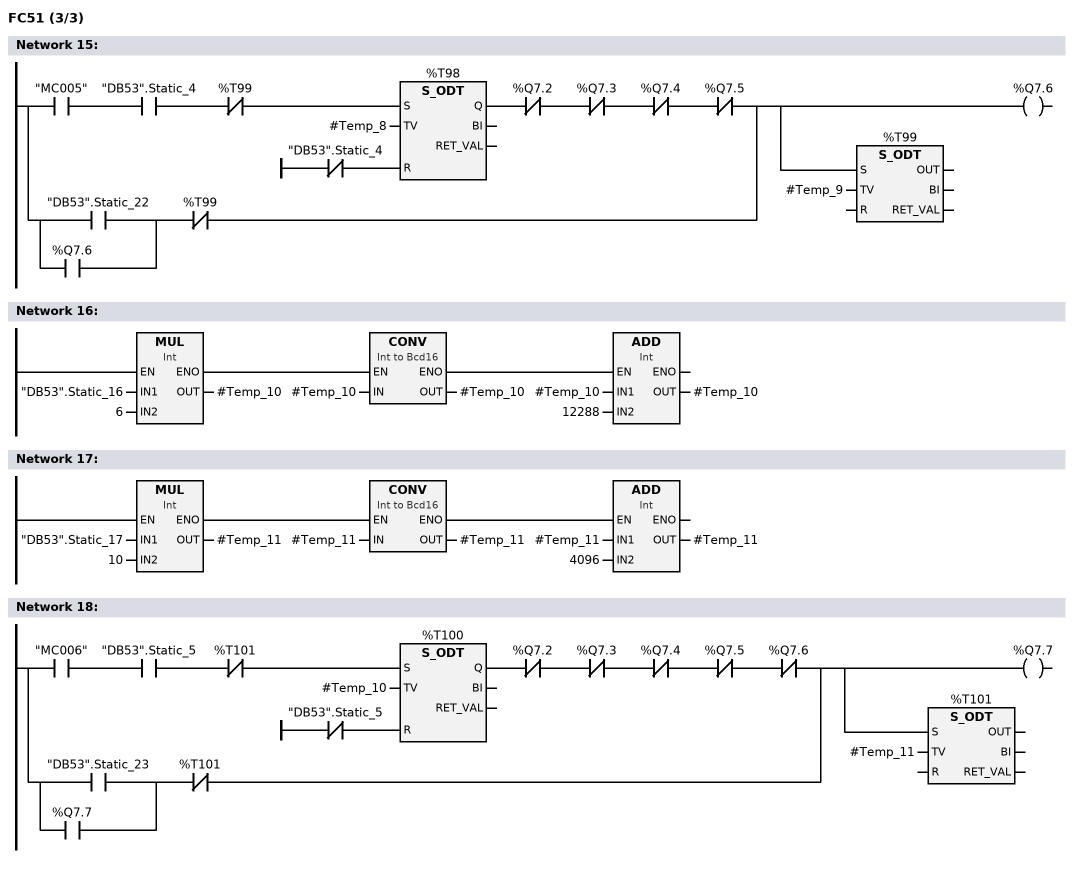
   RUNG wire#powerrail
      Contact( "MC005" )
      Contact( "DB53".Static_4 )
      I_Contact( %T99 )
      S_ODT(T_NO := %T98, TV := #Temp_8, R := wire#w1, BI =>, RET_VAL =>)
      I_Contact( %Q7.2 )
      I_Contact( %Q7.3 )
      I_Contact( %Q7.4 )
      I_Contact( %Q7.5 )
      wire#w2
      Coil( %Q7.6 )
   END_RUNG
   RUNG wire#powerrail
      I_Contact( "DB53".Static_4 )
   END_RUNG wire#w1
   RUNG wire#powerrail
      Contact( "DB53".Static_22 )
      wire#w3
      I_Contact( %T99 )
   END_RUNG wire#w2
   RUNG wire#powerrail
      Contact( %Q7.6 )
   END_RUNG wire#w3
   RUNG wire#w2
      S_ODT(T_NO := %T99, TV := #Temp_9, R :=, BI =>, RET_VAL =>)
   END_RUNG
   // the same network as SCL:
   #_s5time1 := S_ODT(T_NO := %T98,
                      TV := #Temp_8,
                      S := "MC005" AND "DB53".Static_4 AND NOT %T99,
                      R := NOT "DB53".Static_4,
                      Q => #_w1);
   %Q7.6 := (#_w1 AND NOT %Q7.2 AND NOT %Q7.3 AND NOT %Q7.4 AND NOT %Q7.5) OR (("DB53".Static_22 OR %Q7.6) AND NOT %T99);
   #_s5time2 := S_ODT(T_NO := %T99, TV := #Temp_9, S := %Q7.6);
END_REGION

REGION Network 16
   RUNG wire#powerrail
      { S7_Templates := "SrcType := Int"; S7_GenerateENO := "TRUE" } Mul(in1 := "DB53".Static_16, in2 := 6, out => #Temp_10)
      { S7_Templates := "[SrcType := Int, DestType := Bcd16]"; S7_GenerateENO := "TRUE" } Convert(in := #Temp_10, out => #Temp_10)
      { S7_Templates := "SrcType := Int"; S7_GenerateENO := "TRUE" } Add(in1 := #Temp_10, in2 := 12288, out => #Temp_10)
   END_RUNG
   // the same network as SCL:
   // ENO of a box is taken as its EN; it also drops when the box reports an error
   #Temp_10 := "DB53".Static_16 * 6;
   #Temp_10 := INT_TO_BCD16(#Temp_10);
   #Temp_10 := #Temp_10 + 12288;
END_REGION

REGION Network 17
   RUNG wire#powerrail
      { S7_Templates := "SrcType := Int"; S7_GenerateENO := "TRUE" } Mul(in1 := "DB53".Static_17, in2 := 10, out => #Temp_11)
      { S7_Templates := "[SrcType := Int, DestType := Bcd16]"; S7_GenerateENO := "TRUE" } Convert(in := #Temp_11, out => #Temp_11)
      { S7_Templates := "SrcType := Int"; S7_GenerateENO := "TRUE" } Add(in1 := #Temp_11, in2 := 4096, out => #Temp_11)
   END_RUNG
   // the same network as SCL:
   // ENO of a box is taken as its EN; it also drops when the box reports an error
   #Temp_11 := "DB53".Static_17 * 10;
   #Temp_11 := INT_TO_BCD16(#Temp_11);
   #Temp_11 := #Temp_11 + 4096;
END_REGION

REGION Network 18
   RUNG wire#powerrail
      Contact( "MC006" )
      Contact( "DB53".Static_5 )
      I_Contact( %T101 )
      S_ODT(T_NO := %T100, TV := #Temp_10, R := wire#w1, BI =>, RET_VAL =>)
      I_Contact( %Q7.2 )
      I_Contact( %Q7.3 )
      I_Contact( %Q7.4 )
      I_Contact( %Q7.5 )
      I_Contact( %Q7.6 )
      wire#w2
      Coil( %Q7.7 )
   END_RUNG
   RUNG wire#powerrail
      I_Contact( "DB53".Static_5 )
   END_RUNG wire#w1
   RUNG wire#powerrail
      Contact( "DB53".Static_23 )
      wire#w3
      I_Contact( %T101 )
   END_RUNG wire#w2
   RUNG wire#powerrail
      Contact( %Q7.7 )
   END_RUNG wire#w3
   RUNG wire#w2
      S_ODT(T_NO := %T101, TV := #Temp_11, R :=, BI =>, RET_VAL =>)
   END_RUNG
   // the same network as SCL:
   #_s5time1 := S_ODT(T_NO := %T100,
                      TV := #Temp_10,
                      S := "MC006" AND "DB53".Static_5 AND NOT %T101,
                      R := NOT "DB53".Static_5,
                      Q => #_w1);
   %Q7.7 := (#_w1 AND NOT %Q7.2 AND NOT %Q7.3 AND NOT %Q7.4 AND NOT %Q7.5 AND NOT %Q7.6) OR (("DB53".Static_23 OR %Q7.7) AND NOT %T101);
   #_s5time2 := S_ODT(T_NO := %T101, TV := #Temp_11, S := %Q7.7);
END_REGION
END_FUNCTION

ORGANIZATION_BLOCK "Cycle Execution"   // OB1, LAD
{ S7_Optimized_Access := 'FALSE' }
VERSION : 0.1
   VAR_TEMP   // added for the SCL form of the ladder/FBD networks
      _w1 : Bool;
   END_VAR
BEGIN

REGION Network 1
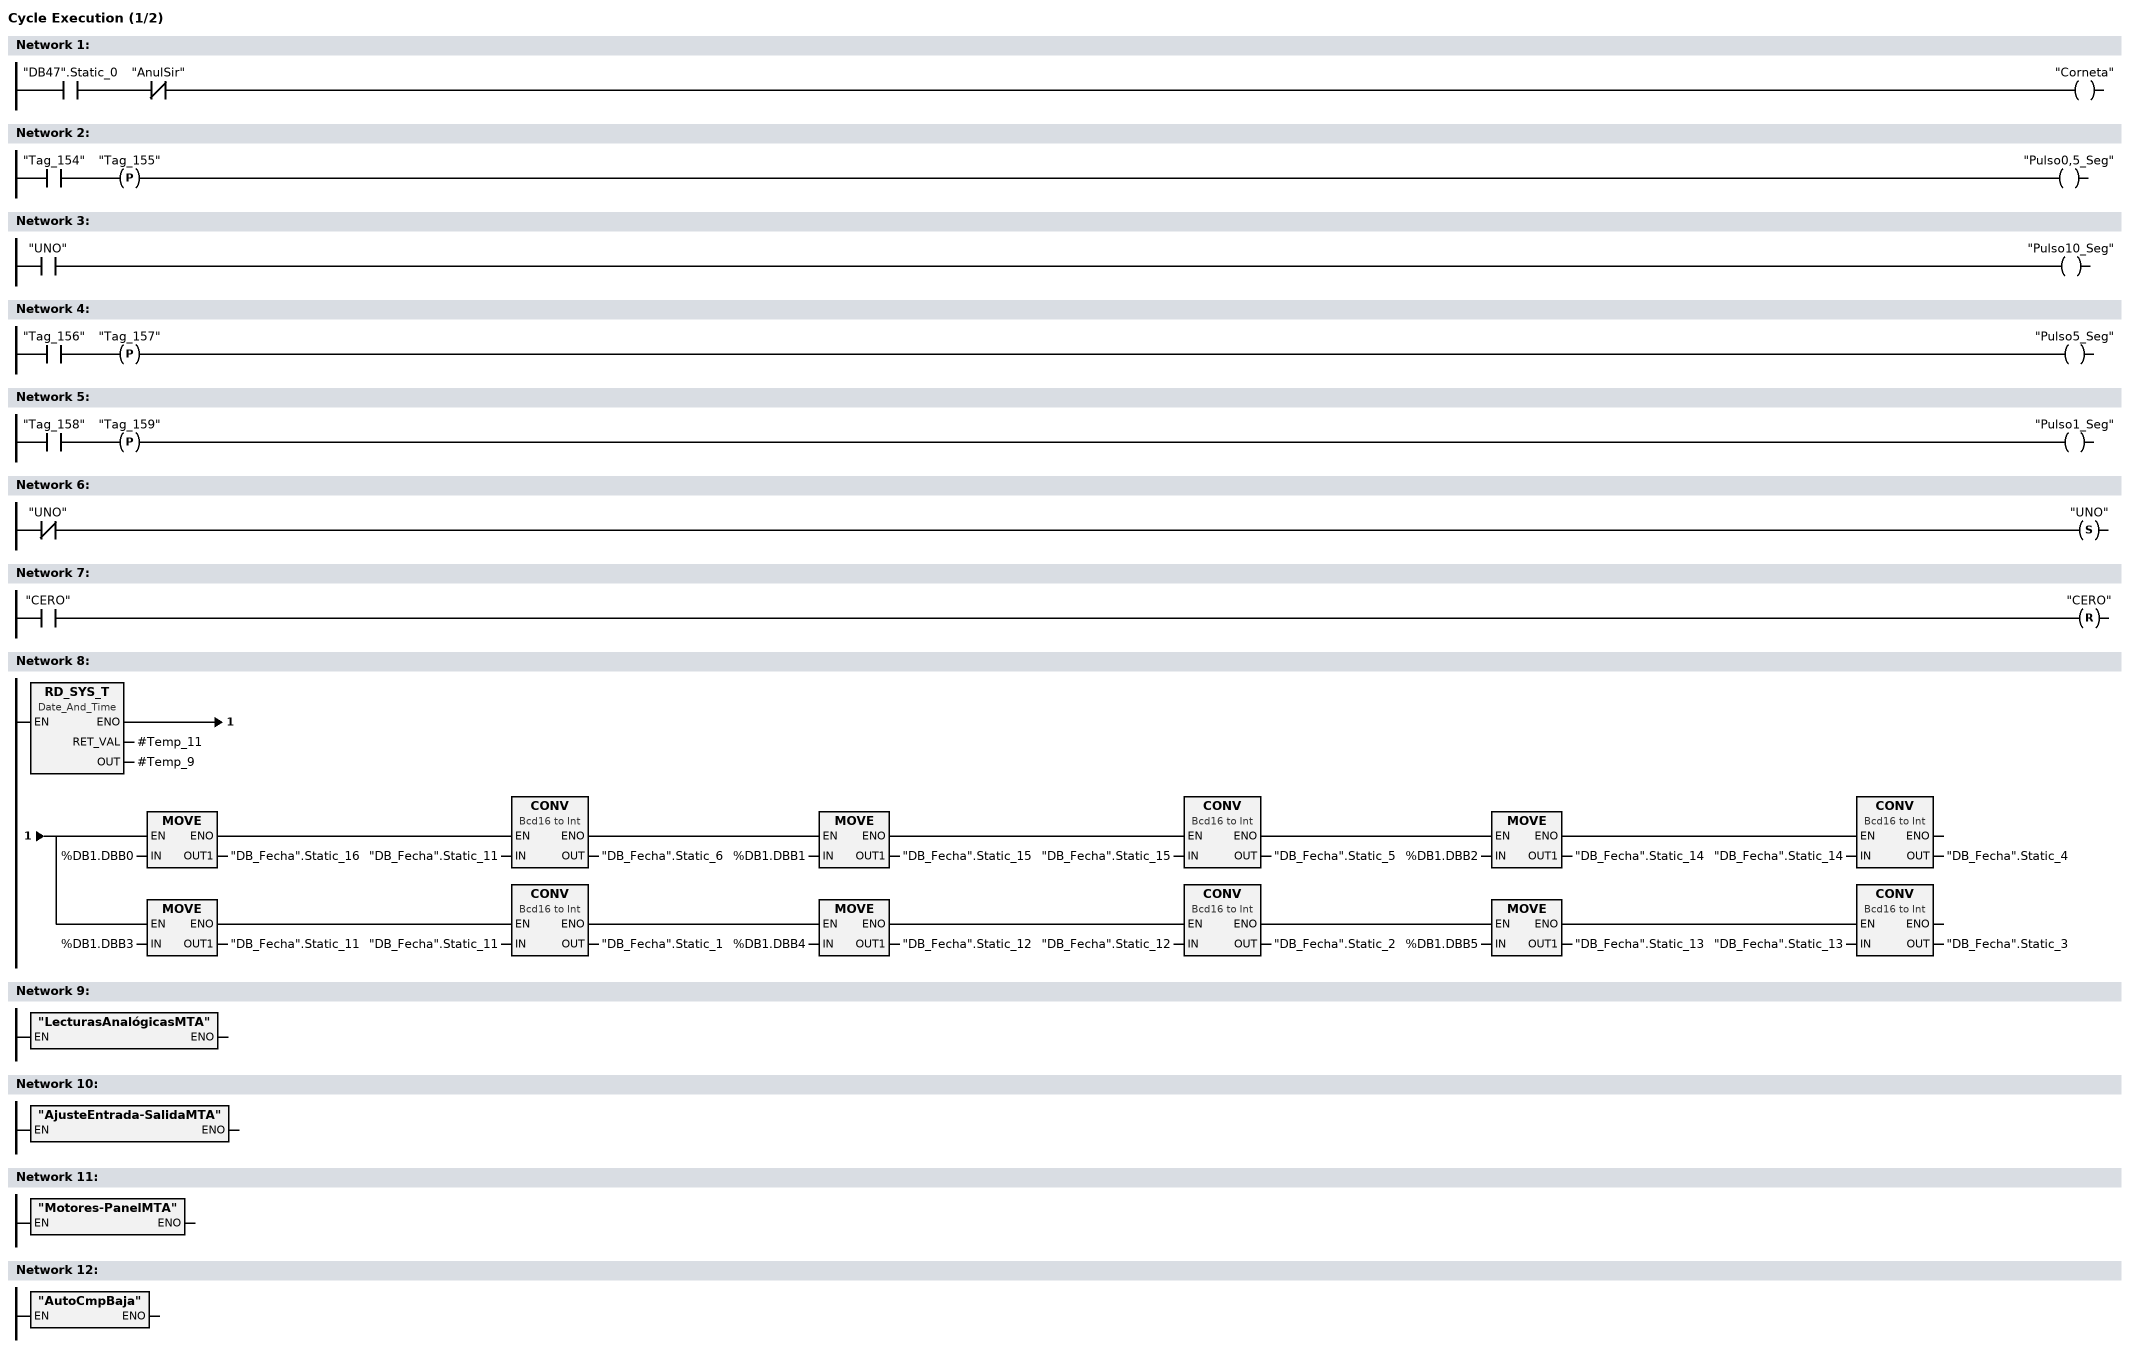
   RUNG wire#powerrail
      Contact( "DB47".Static_0 )
      I_Contact( "AnulSir" )
      Coil( "Corneta" )
   END_RUNG
   // the same network as SCL:
   "Corneta" := "DB47".Static_0 AND NOT "AnulSir";
END_REGION

REGION Network 2
   RUNG wire#powerrail
      Contact( "Tag_154" )
      P_Trig( "Tag_155" )
      Coil( "Pulso0,5_Seg" )
   END_RUNG
   // the same network as SCL:
   #_w1 := "Tag_154" AND NOT "Tag_155";   // rising edge
   "Tag_155" := "Tag_154";
   "Pulso0,5_Seg" := #_w1;
END_REGION

REGION Network 3
   RUNG wire#powerrail
      Contact( "UNO" )
      Coil( "Pulso10_Seg" )
   END_RUNG
   // the same network as SCL:
   "Pulso10_Seg" := "UNO";
END_REGION

REGION Network 4
   RUNG wire#powerrail
      Contact( "Tag_156" )
      P_Trig( "Tag_157" )
      Coil( "Pulso5_Seg" )
   END_RUNG
   // the same network as SCL:
   #_w1 := "Tag_156" AND NOT "Tag_157";   // rising edge
   "Tag_157" := "Tag_156";
   "Pulso5_Seg" := #_w1;
END_REGION

REGION Network 5
   RUNG wire#powerrail
      Contact( "Tag_158" )
      P_Trig( "Tag_159" )
      Coil( "Pulso1_Seg" )
   END_RUNG
   // the same network as SCL:
   #_w1 := "Tag_158" AND NOT "Tag_159";   // rising edge
   "Tag_159" := "Tag_158";
   "Pulso1_Seg" := #_w1;
END_REGION

REGION Network 6
   RUNG wire#powerrail
      I_Contact( "UNO" )
      S_Coil( "UNO" )
   END_RUNG
   // the same network as SCL:
   IF NOT "UNO" THEN "UNO" := TRUE; END_IF;
END_REGION

REGION Network 7
   RUNG wire#powerrail
      Contact( "CERO" )
      R_Coil( "CERO" )
   END_RUNG
   // the same network as SCL:
   IF "CERO" THEN "CERO" := FALSE; END_IF;
END_REGION

REGION Network 8
   // ENO of a box is taken as its EN; it also drops when the box reports an error
   #Temp_11 := RD_SYS_T(out => #Temp_9);
   "DB_Fecha".Static_16 := %DB1.DBB0;
   "DB_Fecha".Static_6 := BCD16_TO_INT("DB_Fecha".Static_11);
   "DB_Fecha".Static_15 := %DB1.DBB1;
   "DB_Fecha".Static_5 := BCD16_TO_INT("DB_Fecha".Static_15);
   "DB_Fecha".Static_14 := %DB1.DBB2;
   "DB_Fecha".Static_4 := BCD16_TO_INT("DB_Fecha".Static_14);
   "DB_Fecha".Static_11 := %DB1.DBB3;
   "DB_Fecha".Static_1 := BCD16_TO_INT("DB_Fecha".Static_11);
   "DB_Fecha".Static_12 := %DB1.DBB4;
   "DB_Fecha".Static_2 := BCD16_TO_INT("DB_Fecha".Static_12);
   "DB_Fecha".Static_13 := %DB1.DBB5;
   "DB_Fecha".Static_3 := BCD16_TO_INT("DB_Fecha".Static_13);
END_REGION

REGION Network 9
   RUNG wire#powerrail
      "LecturasAnalógicasMTA"()
   END_RUNG
   // the same network as SCL:
   "LecturasAnalógicasMTA"();
END_REGION

REGION Network 10
   RUNG wire#powerrail
      "AjusteEntrada-SalidaMTA"()
   END_RUNG
   // the same network as SCL:
   "AjusteEntrada-SalidaMTA"();
END_REGION

REGION Network 11
   RUNG wire#powerrail
      "Motores-PanelMTA"()
   END_RUNG
   // the same network as SCL:
   "Motores-PanelMTA"();
END_REGION

REGION Network 12
   RUNG wire#powerrail
      "AutoCmpBaja"()
   END_RUNG
   // the same network as SCL:
   "AutoCmpBaja"();
END_REGION

REGION Network 13
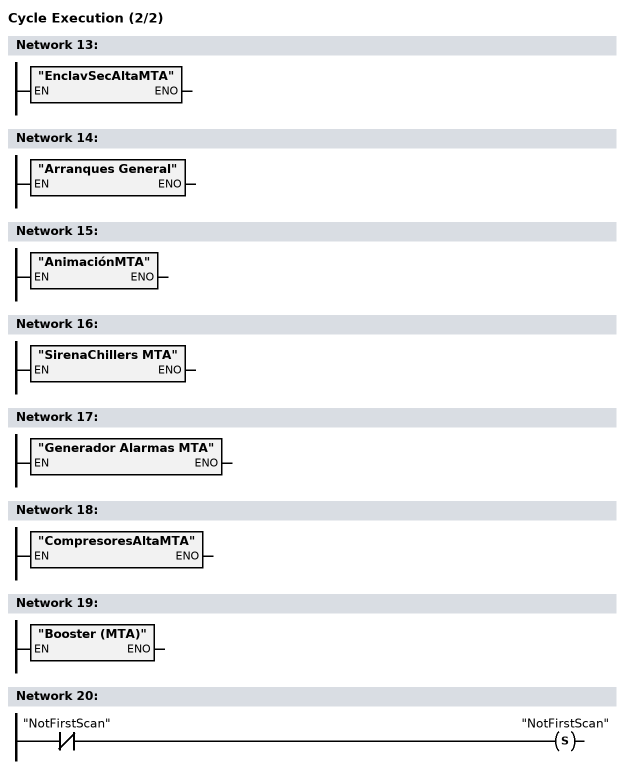
   RUNG wire#powerrail
      "EnclavSecAltaMTA"()
   END_RUNG
   // the same network as SCL:
   "EnclavSecAltaMTA"();
END_REGION

REGION Network 14
   RUNG wire#powerrail
      "Arranques General"()
   END_RUNG
   // the same network as SCL:
   "Arranques General"();
END_REGION

REGION Network 15
   RUNG wire#powerrail
      "AnimaciónMTA"()
   END_RUNG
   // the same network as SCL:
   "AnimaciónMTA"();
END_REGION

REGION Network 16
   RUNG wire#powerrail
      "SirenaChillers MTA"()
   END_RUNG
   // the same network as SCL:
   "SirenaChillers MTA"();
END_REGION

REGION Network 17
   RUNG wire#powerrail
      "Generador Alarmas MTA"()
   END_RUNG
   // the same network as SCL:
   "Generador Alarmas MTA"();
END_REGION

REGION Network 18
   RUNG wire#powerrail
      "CompresoresAltaMTA"()
   END_RUNG
   // the same network as SCL:
   "CompresoresAltaMTA"();
END_REGION

REGION Network 19
   RUNG wire#powerrail
      "Booster (MTA)"()
   END_RUNG
   // the same network as SCL:
   "Booster (MTA)"();
END_REGION

REGION Network 20
   RUNG wire#powerrail
      I_Contact( "NotFirstScan" )
      S_Coil( "NotFirstScan" )
   END_RUNG
   // the same network as SCL:
   IF NOT "NotFirstScan" THEN "NotFirstScan" := TRUE; END_IF;
END_REGION
END_ORGANIZATION_BLOCK

// folder: Alarmas

FUNCTION "SirenaChillers MTA" : Void   // FC7, LAD
{ S7_Optimized_Access := 'FALSE' }
VERSION : 0.1
BEGIN

REGION Network 1
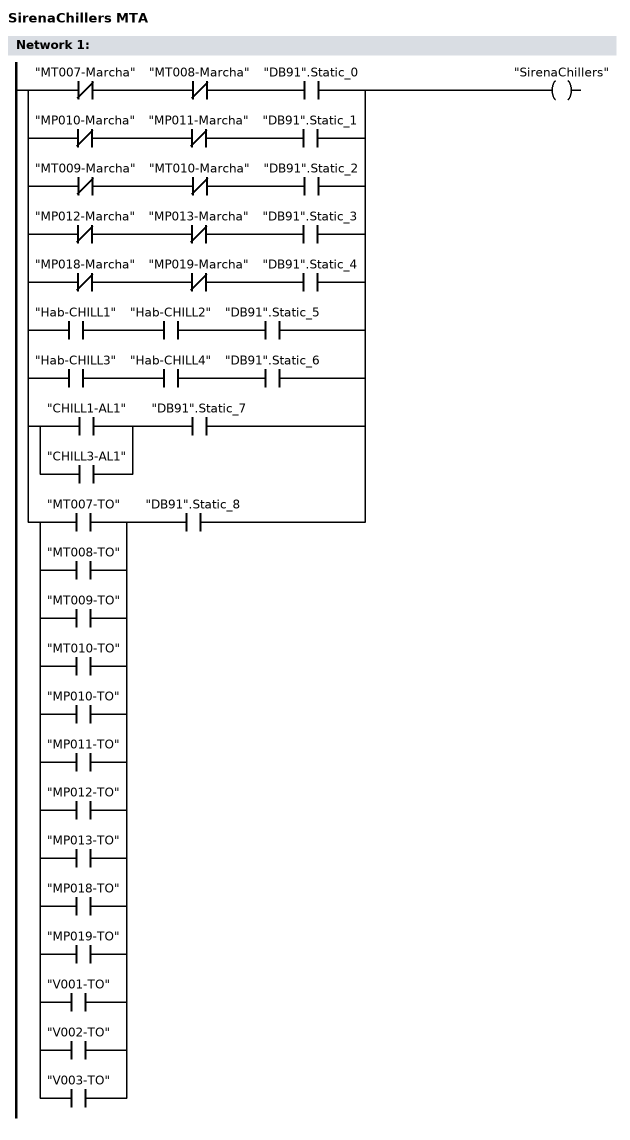
   RUNG wire#powerrail
      I_Contact( "MT007-Marcha" )
      I_Contact( "MT008-Marcha" )
      Contact( "DB91".Static_0 )
      wire#w1
      Coil( "SirenaChillers" )
   END_RUNG
   RUNG wire#powerrail
      I_Contact( "MP010-Marcha" )
      I_Contact( "MP011-Marcha" )
      Contact( "DB91".Static_1 )
   END_RUNG wire#w1
   RUNG wire#powerrail
      I_Contact( "MT009-Marcha" )
      I_Contact( "MT010-Marcha" )
      Contact( "DB91".Static_2 )
   END_RUNG wire#w1
   RUNG wire#powerrail
      I_Contact( "MP012-Marcha" )
      I_Contact( "MP013-Marcha" )
      Contact( "DB91".Static_3 )
   END_RUNG wire#w1
   RUNG wire#powerrail
      I_Contact( "MP018-Marcha" )
      I_Contact( "MP019-Marcha" )
      Contact( "DB91".Static_4 )
   END_RUNG wire#w1
   RUNG wire#powerrail
      Contact( "Hab-CHILL1" )
      Contact( "Hab-CHILL2" )
      Contact( "DB91".Static_5 )
   END_RUNG wire#w1
   RUNG wire#powerrail
      Contact( "Hab-CHILL3" )
      Contact( "Hab-CHILL4" )
      Contact( "DB91".Static_6 )
   END_RUNG wire#w1
   RUNG wire#powerrail
      Contact( "CHILL1-AL1" )
      wire#w2
      Contact( "DB91".Static_7 )
   END_RUNG wire#w1
   RUNG wire#powerrail
      Contact( "CHILL3-AL1" )
   END_RUNG wire#w2
   RUNG wire#powerrail
      Contact( "MT007-TO" )
      wire#w3
      Contact( "DB91".Static_8 )
   END_RUNG wire#w1
   RUNG wire#powerrail
      Contact( "MT008-TO" )
   END_RUNG wire#w3
   RUNG wire#powerrail
      Contact( "MT009-TO" )
   END_RUNG wire#w3
   RUNG wire#powerrail
      Contact( "MT010-TO" )
   END_RUNG wire#w3
   RUNG wire#powerrail
      Contact( "MP010-TO" )
   END_RUNG wire#w3
   RUNG wire#powerrail
      Contact( "MP011-TO" )
   END_RUNG wire#w3
   RUNG wire#powerrail
      Contact( "MP012-TO" )
   END_RUNG wire#w3
   RUNG wire#powerrail
      Contact( "MP013-TO" )
   END_RUNG wire#w3
   RUNG wire#powerrail
      Contact( "MP018-TO" )
   END_RUNG wire#w3
   RUNG wire#powerrail
      Contact( "MP019-TO" )
   END_RUNG wire#w3
   RUNG wire#powerrail
      Contact( "V001-TO" )
   END_RUNG wire#w3
   RUNG wire#powerrail
      Contact( "V002-TO" )
   END_RUNG wire#w3
   RUNG wire#powerrail
      Contact( "V003-TO" )
   END_RUNG wire#w3
   // the same network as SCL:
   "SirenaChillers" := (NOT "MT007-Marcha" AND NOT "MT008-Marcha" AND "DB91".Static_0) OR (NOT "MP010-Marcha" AND NOT "MP011-Marcha" AND "DB91".Static_1) OR (NOT "MT009-Marcha" AND NOT "MT010-Marcha" AND "DB91".Static_2) OR (NOT "MP012-Marcha" AND NOT "MP013-Marcha" AND "DB91".Static_3) OR (NOT "MP018-Marcha" AND NOT "MP019-Marcha" AND "DB91".Static_4) OR ("Hab-CHILL1" AND "Hab-CHILL2" AND "DB91".Static_5) OR ("Hab-CHILL3" AND "Hab-CHILL4" AND "DB91".Static_6) OR (("CHILL1-AL1" OR "CHILL3-AL1") AND "DB91".Static_7) OR (("MT007-TO" OR "MT008-TO" OR "MT009-TO" OR "MT010-TO" OR "MP010-TO" OR "MP011-TO" OR "MP012-TO" OR "MP013-TO" OR "MP018-TO" OR "MP019-TO" OR "V001-TO" OR "V002-TO" OR "V003-TO") AND "DB91".Static_8);
END_REGION
END_FUNCTION

FUNCTION "Generador Alarmas MTA" : Void   // FC8, LAD
{ S7_Optimized_Access := 'FALSE' }
VERSION : 0.1
   VAR_TEMP   // added for the SCL form of the ladder/FBD networks
      _w1 : Bool;
      _s5time1 : S5Time;
   END_VAR
BEGIN

REGION Network 1
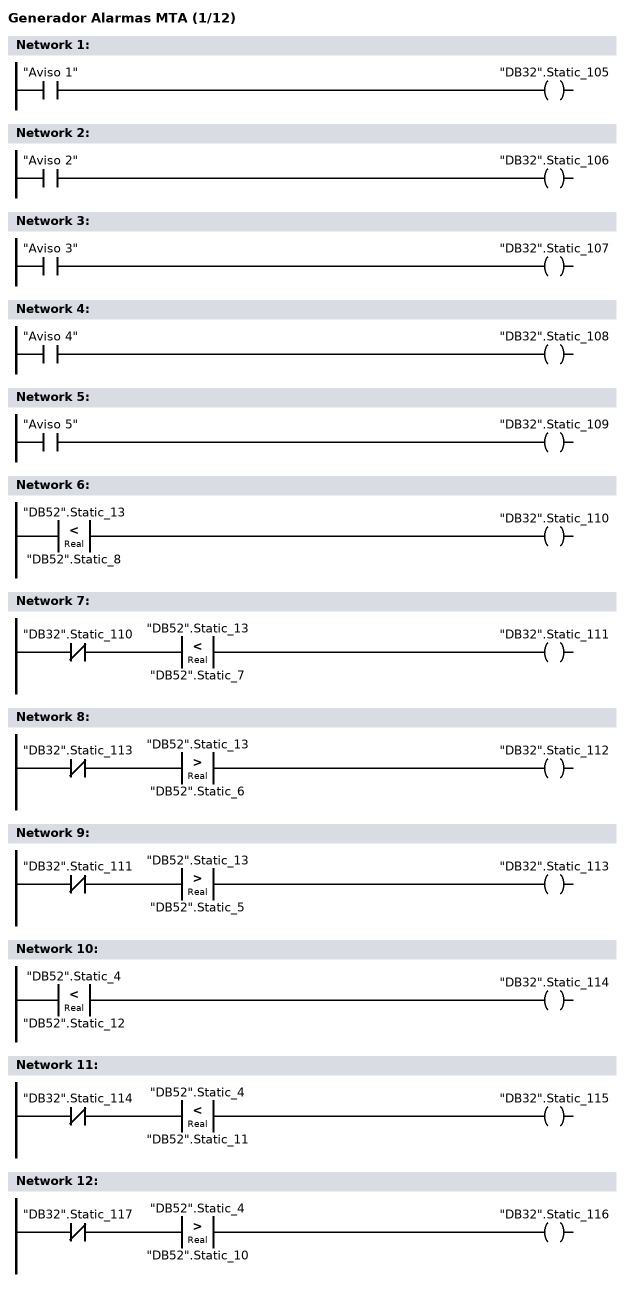
   RUNG wire#powerrail
      Contact( "Aviso 1" )
      Coil( "DB32".Static_105 )
   END_RUNG
   // the same network as SCL:
   "DB32".Static_105 := "Aviso 1";
END_REGION

REGION Network 2
   RUNG wire#powerrail
      Contact( "Aviso 2" )
      Coil( "DB32".Static_106 )
   END_RUNG
   // the same network as SCL:
   "DB32".Static_106 := "Aviso 2";
END_REGION

REGION Network 3
   RUNG wire#powerrail
      Contact( "Aviso 3" )
      Coil( "DB32".Static_107 )
   END_RUNG
   // the same network as SCL:
   "DB32".Static_107 := "Aviso 3";
END_REGION

REGION Network 4
   RUNG wire#powerrail
      Contact( "Aviso 4" )
      Coil( "DB32".Static_108 )
   END_RUNG
   // the same network as SCL:
   "DB32".Static_108 := "Aviso 4";
END_REGION

REGION Network 5
   RUNG wire#powerrail
      Contact( "Aviso 5" )
      Coil( "DB32".Static_109 )
   END_RUNG
   // the same network as SCL:
   "DB32".Static_109 := "Aviso 5";
END_REGION

REGION Network 6
   RUNG wire#powerrail
      { S7_Templates := "SrcType := Real" } LT_Contact(in1 := "DB52".Static_13, in2 := "DB52".Static_8)
      Coil( "DB32".Static_110 )
   END_RUNG
   // the same network as SCL:
   "DB32".Static_110 := "DB52".Static_13 < "DB52".Static_8;
END_REGION

REGION Network 7
   "DB32".Static_111 := NOT "DB32".Static_110 AND ("DB52".Static_13 < "DB52".Static_7);
END_REGION

REGION Network 8
   "DB32".Static_112 := NOT "DB32".Static_113 AND ("DB52".Static_13 > "DB52".Static_6);
END_REGION

REGION Network 9
   "DB32".Static_113 := NOT "DB32".Static_111 AND ("DB52".Static_13 > "DB52".Static_5);
END_REGION

REGION Network 10
   RUNG wire#powerrail
      { S7_Templates := "SrcType := Real" } LT_Contact(in1 := "DB52".Static_4, in2 := "DB52".Static_12)
      Coil( "DB32".Static_114 )
   END_RUNG
   // the same network as SCL:
   "DB32".Static_114 := "DB52".Static_4 < "DB52".Static_12;
END_REGION

REGION Network 11
   "DB32".Static_115 := NOT "DB32".Static_114 AND ("DB52".Static_4 < "DB52".Static_11);
END_REGION

REGION Network 12
   "DB32".Static_116 := NOT "DB32".Static_117 AND ("DB52".Static_4 > "DB52".Static_10);
END_REGION

REGION Network 13
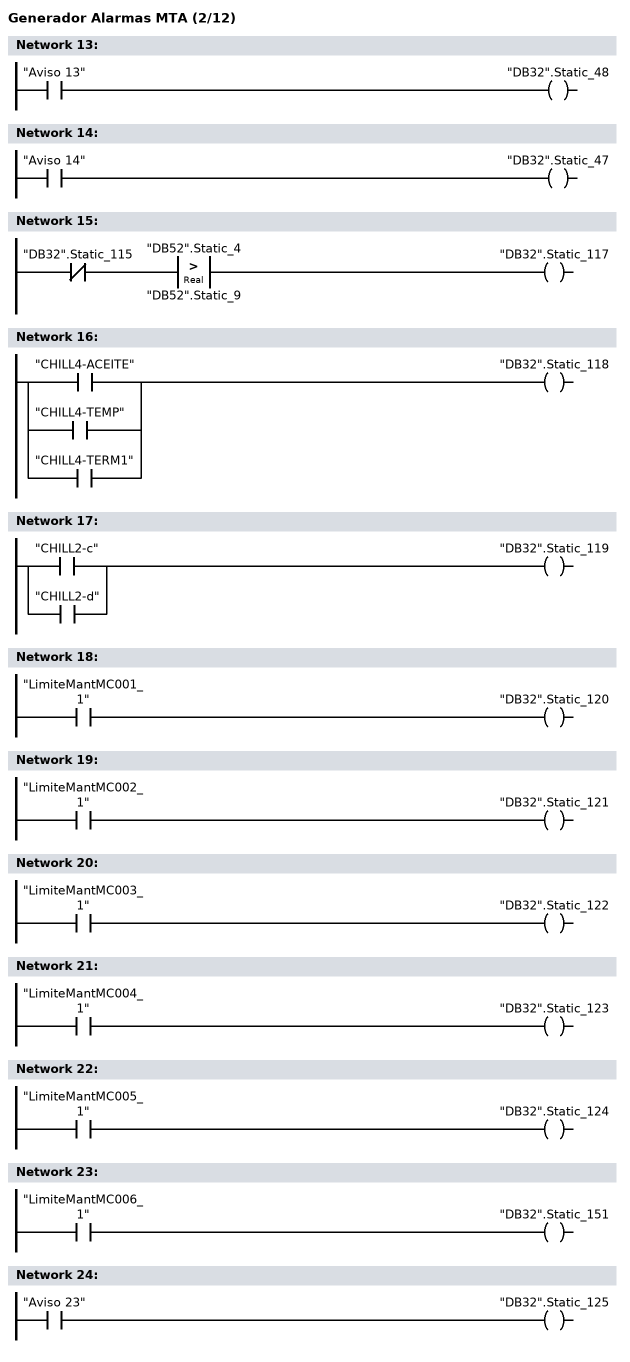
   RUNG wire#powerrail
      Contact( "Aviso 13" )
      Coil( "DB32".Static_48 )
   END_RUNG
   // the same network as SCL:
   "DB32".Static_48 := "Aviso 13";
END_REGION

REGION Network 14
   RUNG wire#powerrail
      Contact( "Aviso 14" )
      Coil( "DB32".Static_47 )
   END_RUNG
   // the same network as SCL:
   "DB32".Static_47 := "Aviso 14";
END_REGION

REGION Network 15
   "DB32".Static_117 := NOT "DB32".Static_115 AND ("DB52".Static_4 > "DB52".Static_9);
END_REGION

REGION Network 16
   RUNG wire#powerrail
      Contact( "CHILL4-ACEITE" )
      wire#w1
      Coil( "DB32".Static_118 )
   END_RUNG
   RUNG wire#powerrail
      Contact( "CHILL4-TEMP" )
   END_RUNG wire#w1
   RUNG wire#powerrail
      Contact( "CHILL4-TERM1" )
   END_RUNG wire#w1
   // the same network as SCL:
   "DB32".Static_118 := "CHILL4-ACEITE" OR "CHILL4-TEMP" OR "CHILL4-TERM1";
END_REGION

REGION Network 17
   RUNG wire#powerrail
      Contact( "CHILL2-c" )
      wire#w1
      Coil( "DB32".Static_119 )
   END_RUNG
   RUNG wire#powerrail
      Contact( "CHILL2-d" )
   END_RUNG wire#w1
   // the same network as SCL:
   "DB32".Static_119 := "CHILL2-c" OR "CHILL2-d";
END_REGION

REGION Network 18
   RUNG wire#powerrail
      Contact( "LimiteMantMC001_1" )
      Coil( "DB32".Static_120 )
   END_RUNG
   // the same network as SCL:
   "DB32".Static_120 := "LimiteMantMC001_1";
END_REGION

REGION Network 19
   RUNG wire#powerrail
      Contact( "LimiteMantMC002_1" )
      Coil( "DB32".Static_121 )
   END_RUNG
   // the same network as SCL:
   "DB32".Static_121 := "LimiteMantMC002_1";
END_REGION

REGION Network 20
   RUNG wire#powerrail
      Contact( "LimiteMantMC003_1" )
      Coil( "DB32".Static_122 )
   END_RUNG
   // the same network as SCL:
   "DB32".Static_122 := "LimiteMantMC003_1";
END_REGION

REGION Network 21
   RUNG wire#powerrail
      Contact( "LimiteMantMC004_1" )
      Coil( "DB32".Static_123 )
   END_RUNG
   // the same network as SCL:
   "DB32".Static_123 := "LimiteMantMC004_1";
END_REGION

REGION Network 22
   RUNG wire#powerrail
      Contact( "LimiteMantMC005_1" )
      Coil( "DB32".Static_124 )
   END_RUNG
   // the same network as SCL:
   "DB32".Static_124 := "LimiteMantMC005_1";
END_REGION

REGION Network 23
   RUNG wire#powerrail
      Contact( "LimiteMantMC006_1" )
      Coil( "DB32".Static_151 )
   END_RUNG
   // the same network as SCL:
   "DB32".Static_151 := "LimiteMantMC006_1";
END_REGION

REGION Network 24
   RUNG wire#powerrail
      Contact( "Aviso 23" )
      Coil( "DB32".Static_125 )
   END_RUNG
   // the same network as SCL:
   "DB32".Static_125 := "Aviso 23";
END_REGION

REGION Network 25
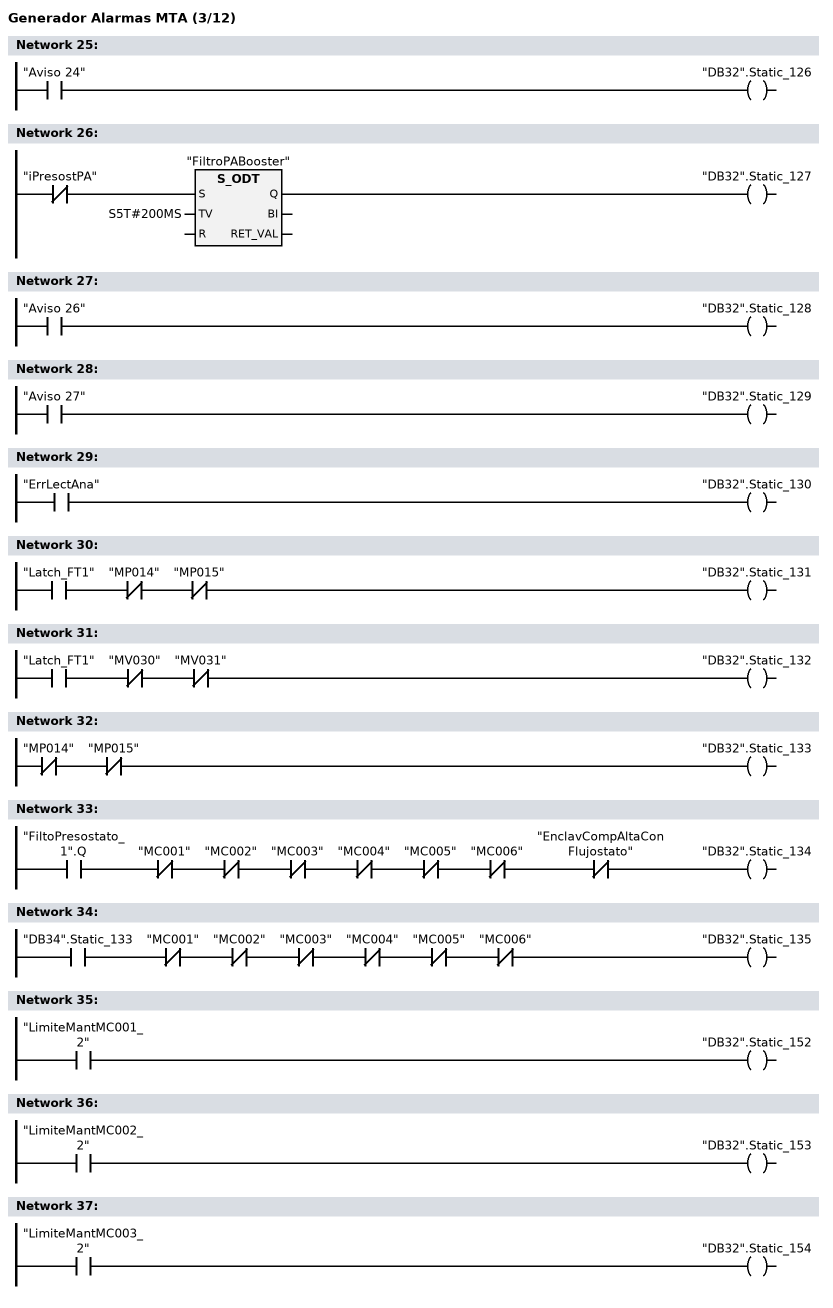
   RUNG wire#powerrail
      Contact( "Aviso 24" )
      Coil( "DB32".Static_126 )
   END_RUNG
   // the same network as SCL:
   "DB32".Static_126 := "Aviso 24";
END_REGION

REGION Network 26
   RUNG wire#powerrail
      I_Contact( "iPresostPA" )
      S_ODT(T_NO := "FiltroPABooster", TV := S5T#200MS, R :=, BI =>, RET_VAL =>)
      Coil( "DB32".Static_127 )
   END_RUNG
   // the same network as SCL:
   #_s5time1 := S_ODT(T_NO := "FiltroPABooster", TV := S5T#200MS, S := NOT "iPresostPA", Q => #_w1);
   "DB32".Static_127 := #_w1;
END_REGION

REGION Network 27
   RUNG wire#powerrail
      Contact( "Aviso 26" )
      Coil( "DB32".Static_128 )
   END_RUNG
   // the same network as SCL:
   "DB32".Static_128 := "Aviso 26";
END_REGION

REGION Network 28
   RUNG wire#powerrail
      Contact( "Aviso 27" )
      Coil( "DB32".Static_129 )
   END_RUNG
   // the same network as SCL:
   "DB32".Static_129 := "Aviso 27";
END_REGION

REGION Network 29
   RUNG wire#powerrail
      Contact( "ErrLectAna" )
      Coil( "DB32".Static_130 )
   END_RUNG
   // the same network as SCL:
   "DB32".Static_130 := "ErrLectAna";
END_REGION

REGION Network 30
   RUNG wire#powerrail
      Contact( "Latch_FT1" )
      I_Contact( "MP014" )
      I_Contact( "MP015" )
      Coil( "DB32".Static_131 )
   END_RUNG
   // the same network as SCL:
   "DB32".Static_131 := "Latch_FT1" AND NOT "MP014" AND NOT "MP015";
END_REGION

REGION Network 31
   RUNG wire#powerrail
      Contact( "Latch_FT1" )
      I_Contact( "MV030" )
      I_Contact( "MV031" )
      Coil( "DB32".Static_132 )
   END_RUNG
   // the same network as SCL:
   "DB32".Static_132 := "Latch_FT1" AND NOT "MV030" AND NOT "MV031";
END_REGION

REGION Network 32
   RUNG wire#powerrail
      I_Contact( "MP014" )
      I_Contact( "MP015" )
      Coil( "DB32".Static_133 )
   END_RUNG
   // the same network as SCL:
   "DB32".Static_133 := NOT "MP014" AND NOT "MP015";
END_REGION

REGION Network 33
   RUNG wire#powerrail
      Contact( "FiltoPresostato_1".Q )
      I_Contact( "MC001" )
      I_Contact( "MC002" )
      I_Contact( "MC003" )
      I_Contact( "MC004" )
      I_Contact( "MC005" )
      I_Contact( "MC006" )
      I_Contact( "EnclavCompAltaConFlujostato" )
      Coil( "DB32".Static_134 )
   END_RUNG
   // the same network as SCL:
   "DB32".Static_134 := "FiltoPresostato_1".Q AND NOT "MC001" AND NOT "MC002" AND NOT "MC003" AND NOT "MC004" AND NOT "MC005" AND NOT "MC006" AND NOT "EnclavCompAltaConFlujostato";
END_REGION

REGION Network 34
   RUNG wire#powerrail
      Contact( "DB34".Static_133 )
      I_Contact( "MC001" )
      I_Contact( "MC002" )
      I_Contact( "MC003" )
      I_Contact( "MC004" )
      I_Contact( "MC005" )
      I_Contact( "MC006" )
      Coil( "DB32".Static_135 )
   END_RUNG
   // the same network as SCL:
   "DB32".Static_135 := "DB34".Static_133 AND NOT "MC001" AND NOT "MC002" AND NOT "MC003" AND NOT "MC004" AND NOT "MC005" AND NOT "MC006";
END_REGION

REGION Network 35
   RUNG wire#powerrail
      Contact( "LimiteMantMC001_2" )
      Coil( "DB32".Static_152 )
   END_RUNG
   // the same network as SCL:
   "DB32".Static_152 := "LimiteMantMC001_2";
END_REGION

REGION Network 36
   RUNG wire#powerrail
      Contact( "LimiteMantMC002_2" )
      Coil( "DB32".Static_153 )
   END_RUNG
   // the same network as SCL:
   "DB32".Static_153 := "LimiteMantMC002_2";
END_REGION

REGION Network 37
   RUNG wire#powerrail
      Contact( "LimiteMantMC003_2" )
      Coil( "DB32".Static_154 )
   END_RUNG
   // the same network as SCL:
   "DB32".Static_154 := "LimiteMantMC003_2";
END_REGION

REGION Network 38
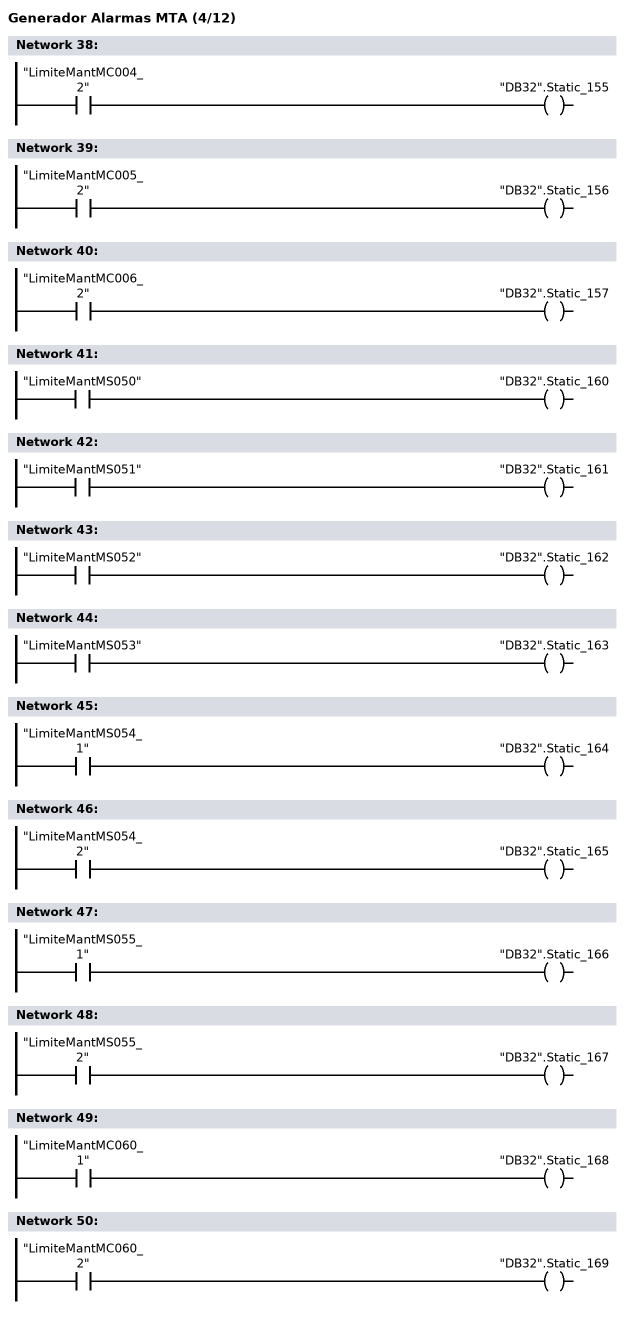
   RUNG wire#powerrail
      Contact( "LimiteMantMC004_2" )
      Coil( "DB32".Static_155 )
   END_RUNG
   // the same network as SCL:
   "DB32".Static_155 := "LimiteMantMC004_2";
END_REGION

REGION Network 39
   RUNG wire#powerrail
      Contact( "LimiteMantMC005_2" )
      Coil( "DB32".Static_156 )
   END_RUNG
   // the same network as SCL:
   "DB32".Static_156 := "LimiteMantMC005_2";
END_REGION

REGION Network 40
   RUNG wire#powerrail
      Contact( "LimiteMantMC006_2" )
      Coil( "DB32".Static_157 )
   END_RUNG
   // the same network as SCL:
   "DB32".Static_157 := "LimiteMantMC006_2";
END_REGION

REGION Network 41
   RUNG wire#powerrail
      Contact( "LimiteMantMS050" )
      Coil( "DB32".Static_160 )
   END_RUNG
   // the same network as SCL:
   "DB32".Static_160 := "LimiteMantMS050";
END_REGION

REGION Network 42
   RUNG wire#powerrail
      Contact( "LimiteMantMS051" )
      Coil( "DB32".Static_161 )
   END_RUNG
   // the same network as SCL:
   "DB32".Static_161 := "LimiteMantMS051";
END_REGION

REGION Network 43
   RUNG wire#powerrail
      Contact( "LimiteMantMS052" )
      Coil( "DB32".Static_162 )
   END_RUNG
   // the same network as SCL:
   "DB32".Static_162 := "LimiteMantMS052";
END_REGION

REGION Network 44
   RUNG wire#powerrail
      Contact( "LimiteMantMS053" )
      Coil( "DB32".Static_163 )
   END_RUNG
   // the same network as SCL:
   "DB32".Static_163 := "LimiteMantMS053";
END_REGION

REGION Network 45
   RUNG wire#powerrail
      Contact( "LimiteMantMS054_1" )
      Coil( "DB32".Static_164 )
   END_RUNG
   // the same network as SCL:
   "DB32".Static_164 := "LimiteMantMS054_1";
END_REGION

REGION Network 46
   RUNG wire#powerrail
      Contact( "LimiteMantMS054_2" )
      Coil( "DB32".Static_165 )
   END_RUNG
   // the same network as SCL:
   "DB32".Static_165 := "LimiteMantMS054_2";
END_REGION

REGION Network 47
   RUNG wire#powerrail
      Contact( "LimiteMantMS055_1" )
      Coil( "DB32".Static_166 )
   END_RUNG
   // the same network as SCL:
   "DB32".Static_166 := "LimiteMantMS055_1";
END_REGION

REGION Network 48
   RUNG wire#powerrail
      Contact( "LimiteMantMS055_2" )
      Coil( "DB32".Static_167 )
   END_RUNG
   // the same network as SCL:
   "DB32".Static_167 := "LimiteMantMS055_2";
END_REGION

REGION Network 49
   RUNG wire#powerrail
      Contact( "LimiteMantMC060_1" )
      Coil( "DB32".Static_168 )
   END_RUNG
   // the same network as SCL:
   "DB32".Static_168 := "LimiteMantMC060_1";
END_REGION

REGION Network 50
   RUNG wire#powerrail
      Contact( "LimiteMantMC060_2" )
      Coil( "DB32".Static_169 )
   END_RUNG
   // the same network as SCL:
   "DB32".Static_169 := "LimiteMantMC060_2";
END_REGION

REGION Network 51
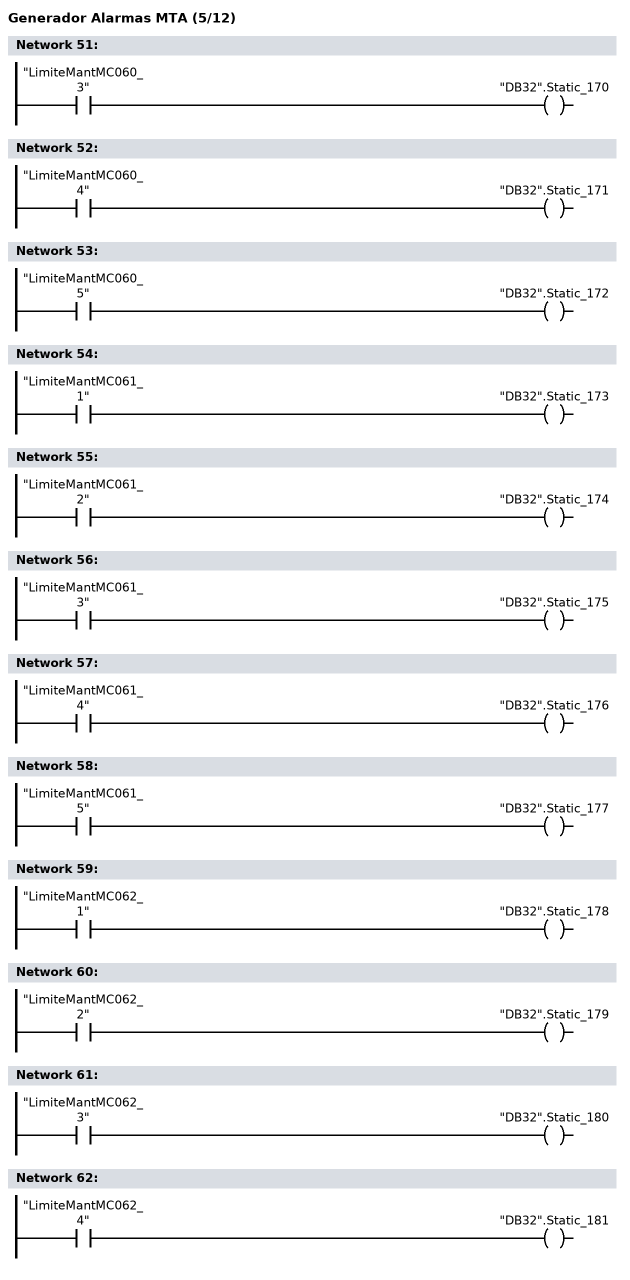
   RUNG wire#powerrail
      Contact( "LimiteMantMC060_3" )
      Coil( "DB32".Static_170 )
   END_RUNG
   // the same network as SCL:
   "DB32".Static_170 := "LimiteMantMC060_3";
END_REGION

REGION Network 52
   RUNG wire#powerrail
      Contact( "LimiteMantMC060_4" )
      Coil( "DB32".Static_171 )
   END_RUNG
   // the same network as SCL:
   "DB32".Static_171 := "LimiteMantMC060_4";
END_REGION

REGION Network 53
   RUNG wire#powerrail
      Contact( "LimiteMantMC060_5" )
      Coil( "DB32".Static_172 )
   END_RUNG
   // the same network as SCL:
   "DB32".Static_172 := "LimiteMantMC060_5";
END_REGION

REGION Network 54
   RUNG wire#powerrail
      Contact( "LimiteMantMC061_1" )
      Coil( "DB32".Static_173 )
   END_RUNG
   // the same network as SCL:
   "DB32".Static_173 := "LimiteMantMC061_1";
END_REGION

REGION Network 55
   RUNG wire#powerrail
      Contact( "LimiteMantMC061_2" )
      Coil( "DB32".Static_174 )
   END_RUNG
   // the same network as SCL:
   "DB32".Static_174 := "LimiteMantMC061_2";
END_REGION

REGION Network 56
   RUNG wire#powerrail
      Contact( "LimiteMantMC061_3" )
      Coil( "DB32".Static_175 )
   END_RUNG
   // the same network as SCL:
   "DB32".Static_175 := "LimiteMantMC061_3";
END_REGION

REGION Network 57
   RUNG wire#powerrail
      Contact( "LimiteMantMC061_4" )
      Coil( "DB32".Static_176 )
   END_RUNG
   // the same network as SCL:
   "DB32".Static_176 := "LimiteMantMC061_4";
END_REGION

REGION Network 58
   RUNG wire#powerrail
      Contact( "LimiteMantMC061_5" )
      Coil( "DB32".Static_177 )
   END_RUNG
   // the same network as SCL:
   "DB32".Static_177 := "LimiteMantMC061_5";
END_REGION

REGION Network 59
   RUNG wire#powerrail
      Contact( "LimiteMantMC062_1" )
      Coil( "DB32".Static_178 )
   END_RUNG
   // the same network as SCL:
   "DB32".Static_178 := "LimiteMantMC062_1";
END_REGION

REGION Network 60
   RUNG wire#powerrail
      Contact( "LimiteMantMC062_2" )
      Coil( "DB32".Static_179 )
   END_RUNG
   // the same network as SCL:
   "DB32".Static_179 := "LimiteMantMC062_2";
END_REGION

REGION Network 61
   RUNG wire#powerrail
      Contact( "LimiteMantMC062_3" )
      Coil( "DB32".Static_180 )
   END_RUNG
   // the same network as SCL:
   "DB32".Static_180 := "LimiteMantMC062_3";
END_REGION

REGION Network 62
   RUNG wire#powerrail
      Contact( "LimiteMantMC062_4" )
      Coil( "DB32".Static_181 )
   END_RUNG
   // the same network as SCL:
   "DB32".Static_181 := "LimiteMantMC062_4";
END_REGION

REGION Network 63
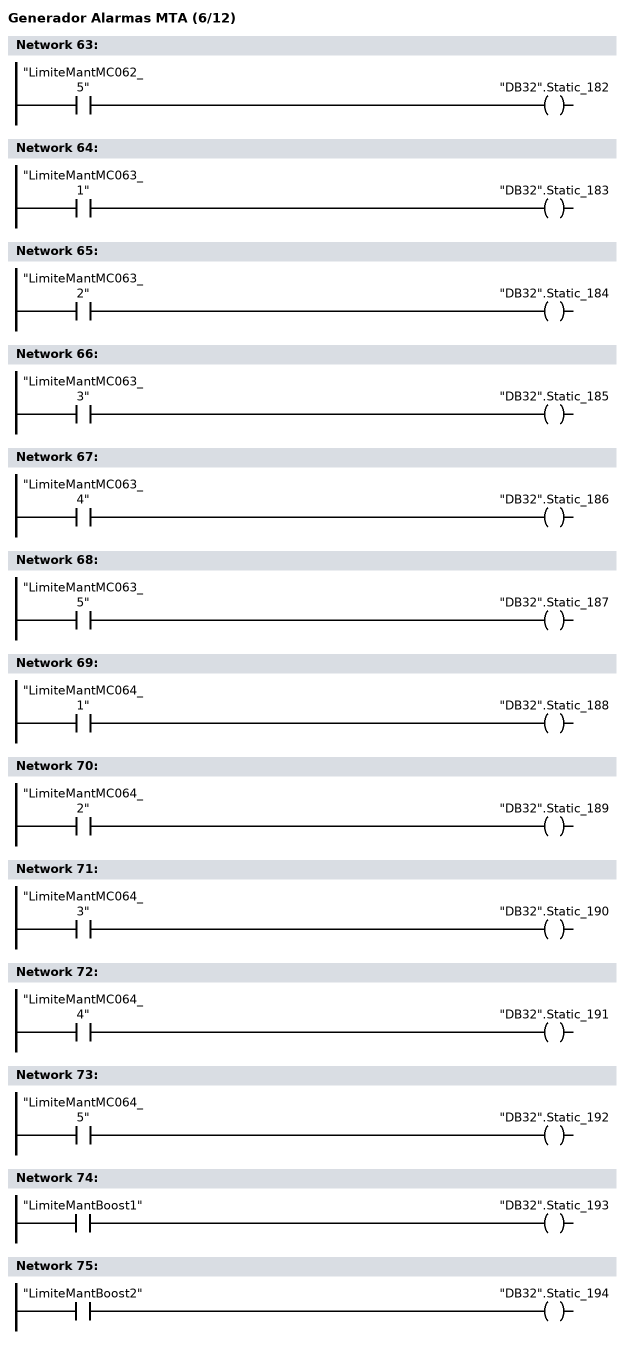
   RUNG wire#powerrail
      Contact( "LimiteMantMC062_5" )
      Coil( "DB32".Static_182 )
   END_RUNG
   // the same network as SCL:
   "DB32".Static_182 := "LimiteMantMC062_5";
END_REGION

REGION Network 64
   RUNG wire#powerrail
      Contact( "LimiteMantMC063_1" )
      Coil( "DB32".Static_183 )
   END_RUNG
   // the same network as SCL:
   "DB32".Static_183 := "LimiteMantMC063_1";
END_REGION

REGION Network 65
   RUNG wire#powerrail
      Contact( "LimiteMantMC063_2" )
      Coil( "DB32".Static_184 )
   END_RUNG
   // the same network as SCL:
   "DB32".Static_184 := "LimiteMantMC063_2";
END_REGION

REGION Network 66
   RUNG wire#powerrail
      Contact( "LimiteMantMC063_3" )
      Coil( "DB32".Static_185 )
   END_RUNG
   // the same network as SCL:
   "DB32".Static_185 := "LimiteMantMC063_3";
END_REGION

REGION Network 67
   RUNG wire#powerrail
      Contact( "LimiteMantMC063_4" )
      Coil( "DB32".Static_186 )
   END_RUNG
   // the same network as SCL:
   "DB32".Static_186 := "LimiteMantMC063_4";
END_REGION

REGION Network 68
   RUNG wire#powerrail
      Contact( "LimiteMantMC063_5" )
      Coil( "DB32".Static_187 )
   END_RUNG
   // the same network as SCL:
   "DB32".Static_187 := "LimiteMantMC063_5";
END_REGION

REGION Network 69
   RUNG wire#powerrail
      Contact( "LimiteMantMC064_1" )
      Coil( "DB32".Static_188 )
   END_RUNG
   // the same network as SCL:
   "DB32".Static_188 := "LimiteMantMC064_1";
END_REGION

REGION Network 70
   RUNG wire#powerrail
      Contact( "LimiteMantMC064_2" )
      Coil( "DB32".Static_189 )
   END_RUNG
   // the same network as SCL:
   "DB32".Static_189 := "LimiteMantMC064_2";
END_REGION

REGION Network 71
   RUNG wire#powerrail
      Contact( "LimiteMantMC064_3" )
      Coil( "DB32".Static_190 )
   END_RUNG
   // the same network as SCL:
   "DB32".Static_190 := "LimiteMantMC064_3";
END_REGION

REGION Network 72
   RUNG wire#powerrail
      Contact( "LimiteMantMC064_4" )
      Coil( "DB32".Static_191 )
   END_RUNG
   // the same network as SCL:
   "DB32".Static_191 := "LimiteMantMC064_4";
END_REGION

REGION Network 73
   RUNG wire#powerrail
      Contact( "LimiteMantMC064_5" )
      Coil( "DB32".Static_192 )
   END_RUNG
   // the same network as SCL:
   "DB32".Static_192 := "LimiteMantMC064_5";
END_REGION

REGION Network 74
   RUNG wire#powerrail
      Contact( "LimiteMantBoost1" )
      Coil( "DB32".Static_193 )
   END_RUNG
   // the same network as SCL:
   "DB32".Static_193 := "LimiteMantBoost1";
END_REGION

